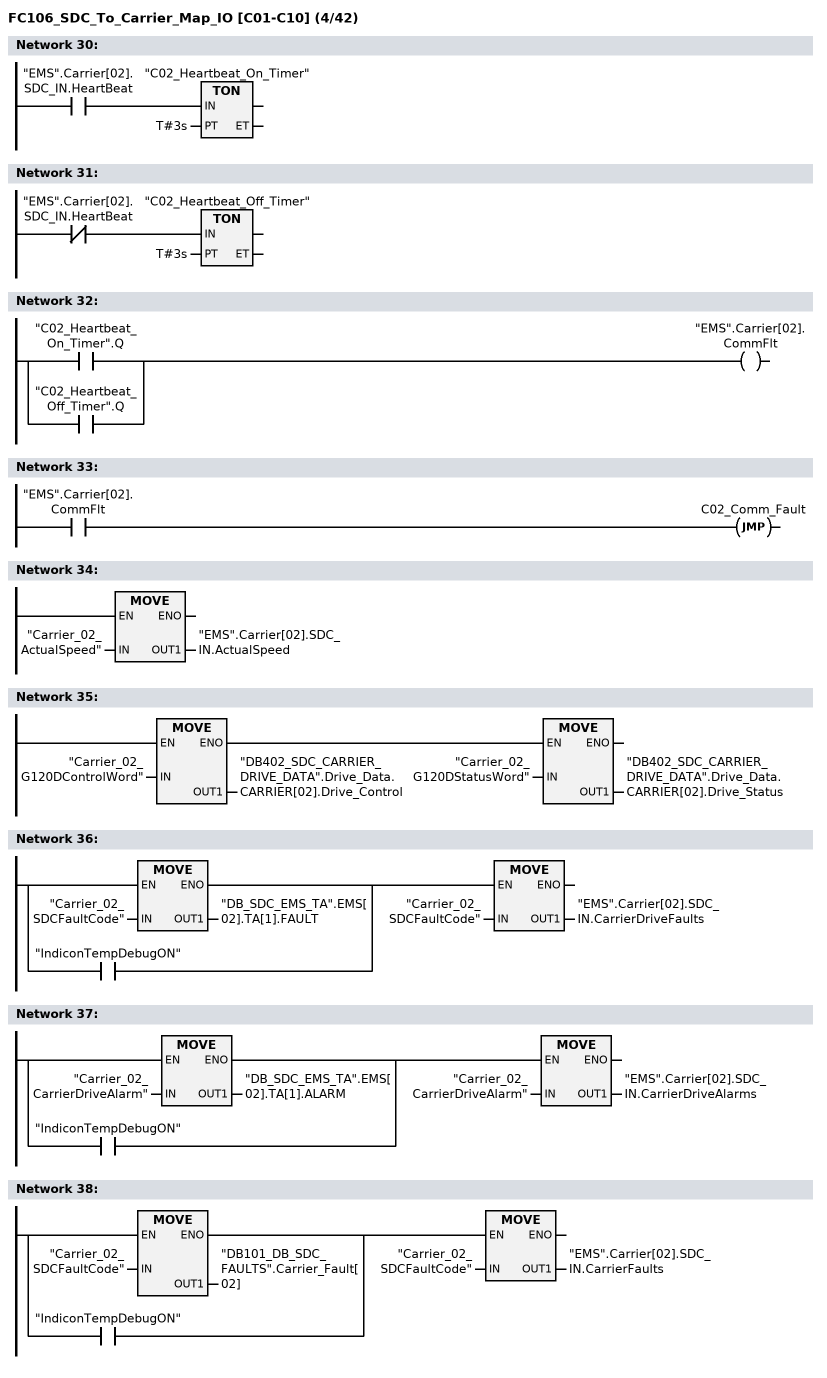
   "C02_Heartbeat_On_Timer".TON(IN := "EMS".Carrier[02].SDC_IN.HeartBeat, PT := T#3s);
END_REGION

REGION Network 31
   "C02_Heartbeat_Off_Timer".TON(IN := NOT "EMS".Carrier[02].SDC_IN.HeartBeat, PT := T#3s);
END_REGION

REGION Network 32
   RUNG wire#powerrail
      Contact( "C02_Heartbeat_On_Timer".Q )
      wire#w1
      Coil( "EMS".Carrier[02].CommFlt )
   END_RUNG
   RUNG wire#powerrail
      Contact( "C02_Heartbeat_Off_Timer".Q )
   END_RUNG wire#w1
   // the same network as SCL:
   "EMS".Carrier[02].CommFlt := "C02_Heartbeat_On_Timer".Q OR "C02_Heartbeat_Off_Timer".Q;
END_REGION

REGION Network 33
   RUNG wire#powerrail
      Contact( "EMS".Carrier[02].CommFlt )
      JumpCoil( C02_Comm_Fault )
   END_RUNG
   // the same network as SCL:
   IF "EMS".Carrier[02].CommFlt THEN GOTO C02_Comm_Fault; END_IF;
END_REGION

REGION Network 34
   RUNG wire#powerrail
      Move(in := "Carrier_02_ActualSpeed", out1 => "EMS".Carrier[02].SDC_IN.ActualSpeed)
   END_RUNG
   // the same network as SCL:
   "EMS".Carrier[02].SDC_IN.ActualSpeed := "Carrier_02_ActualSpeed";
END_REGION

REGION Network 35
   RUNG wire#powerrail
      Move(in := "Carrier_02_G120DControlWord", out1 => "DB402_SDC_CARRIER_DRIVE_DATA".Drive_Data.CARRIER[02].Drive_Control)
      Move(in := "Carrier_02_G120DStatusWord", out1 => "DB402_SDC_CARRIER_DRIVE_DATA".Drive_Data.CARRIER[02].Drive_Status)
   END_RUNG
   // the same network as SCL:
   "DB402_SDC_CARRIER_DRIVE_DATA".Drive_Data.CARRIER[02].Drive_Control := "Carrier_02_G120DControlWord";
   "DB402_SDC_CARRIER_DRIVE_DATA".Drive_Data.CARRIER[02].Drive_Status := "Carrier_02_G120DStatusWord";
END_REGION

REGION Network 36
   RUNG wire#powerrail
      Move(in := "Carrier_02_SDCFaultCode", out1 => "DB_SDC_EMS_TA".EMS[02].TA[1].FAULT)
      wire#w1
      Move(in := "Carrier_02_SDCFaultCode", out1 => "EMS".Carrier[02].SDC_IN.CarrierDriveFaults)
   END_RUNG
   RUNG wire#powerrail
      Contact( "IndiconTempDebugON" )
   END_RUNG wire#w1
   // the same network as SCL:
   "DB_SDC_EMS_TA".EMS[02].TA[1].FAULT := "Carrier_02_SDCFaultCode";
   IF TRUE OR "IndiconTempDebugON" THEN
       "EMS".Carrier[02].SDC_IN.CarrierDriveFaults := "Carrier_02_SDCFaultCode";
   END_IF;
END_REGION

REGION Network 37
   RUNG wire#powerrail
      Move(in := "Carrier_02_CarrierDriveAlarm", out1 => "DB_SDC_EMS_TA".EMS[02].TA[1].ALARM)
      wire#w1
      Move(in := "Carrier_02_CarrierDriveAlarm", out1 => "EMS".Carrier[02].SDC_IN.CarrierDriveAlarms)
   END_RUNG
   RUNG wire#powerrail
      Contact( "IndiconTempDebugON" )
   END_RUNG wire#w1
   // the same network as SCL:
   "DB_SDC_EMS_TA".EMS[02].TA[1].ALARM := "Carrier_02_CarrierDriveAlarm";
   IF TRUE OR "IndiconTempDebugON" THEN
       "EMS".Carrier[02].SDC_IN.CarrierDriveAlarms := "Carrier_02_CarrierDriveAlarm";
   END_IF;
END_REGION

REGION Network 38
   RUNG wire#powerrail
      Move(in := "Carrier_02_SDCFaultCode", out1 => "DB101_DB_SDC_FAULTS".Carrier_Fault[02])
      wire#w1
      Move(in := "Carrier_02_SDCFaultCode", out1 => "EMS".Carrier[02].SDC_IN.CarrierFaults)
   END_RUNG
   RUNG wire#powerrail
      Contact( "IndiconTempDebugON" )
   END_RUNG wire#w1
   // the same network as SCL:
   "DB101_DB_SDC_FAULTS".Carrier_Fault[02] := "Carrier_02_SDCFaultCode";
   IF TRUE OR "IndiconTempDebugON" THEN
       "EMS".Carrier[02].SDC_IN.CarrierFaults := "Carrier_02_SDCFaultCode";
   END_IF;
END_REGION

REGION Network 39
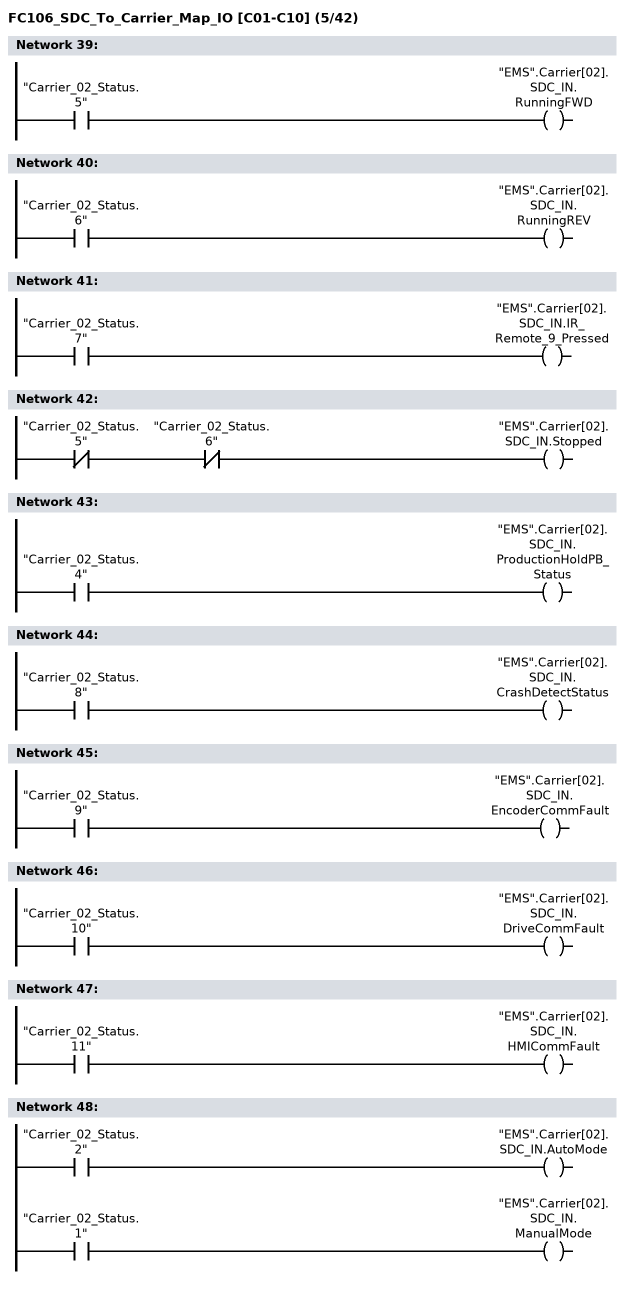
   RUNG wire#powerrail
      Contact( "Carrier_02_Status.5" )
      Coil( "EMS".Carrier[02].SDC_IN.RunningFWD )
   END_RUNG
   // the same network as SCL:
   "EMS".Carrier[02].SDC_IN.RunningFWD := "Carrier_02_Status.5";
END_REGION

REGION Network 40
   RUNG wire#powerrail
      Contact( "Carrier_02_Status.6" )
      Coil( "EMS".Carrier[02].SDC_IN.RunningREV )
   END_RUNG
   // the same network as SCL:
   "EMS".Carrier[02].SDC_IN.RunningREV := "Carrier_02_Status.6";
END_REGION

REGION Network 41
   RUNG wire#powerrail
      Contact( "Carrier_02_Status.7" )
      Coil( "EMS".Carrier[02].SDC_IN.IR_Remote_9_Pressed )
   END_RUNG
   // the same network as SCL:
   "EMS".Carrier[02].SDC_IN.IR_Remote_9_Pressed := "Carrier_02_Status.7";
END_REGION

REGION Network 42
   RUNG wire#powerrail
      I_Contact( "Carrier_02_Status.5" )
      I_Contact( "Carrier_02_Status.6" )
      Coil( "EMS".Carrier[02].SDC_IN.Stopped )
   END_RUNG
   // the same network as SCL:
   "EMS".Carrier[02].SDC_IN.Stopped := NOT "Carrier_02_Status.5" AND NOT "Carrier_02_Status.6";
END_REGION

REGION Network 43
   RUNG wire#powerrail
      Contact( "Carrier_02_Status.4" )
      Coil( "EMS".Carrier[02].SDC_IN.ProductionHoldPB_Status )
   END_RUNG
   // the same network as SCL:
   "EMS".Carrier[02].SDC_IN.ProductionHoldPB_Status := "Carrier_02_Status.4";
END_REGION

REGION Network 44
   RUNG wire#powerrail
      Contact( "Carrier_02_Status.8" )
      Coil( "EMS".Carrier[02].SDC_IN.CrashDetectStatus )
   END_RUNG
   // the same network as SCL:
   "EMS".Carrier[02].SDC_IN.CrashDetectStatus := "Carrier_02_Status.8";
END_REGION

REGION Network 45
   RUNG wire#powerrail
      Contact( "Carrier_02_Status.9" )
      Coil( "EMS".Carrier[02].SDC_IN.EncoderCommFault )
   END_RUNG
   // the same network as SCL:
   "EMS".Carrier[02].SDC_IN.EncoderCommFault := "Carrier_02_Status.9";
END_REGION

REGION Network 46
   RUNG wire#powerrail
      Contact( "Carrier_02_Status.10" )
      Coil( "EMS".Carrier[02].SDC_IN.DriveCommFault )
   END_RUNG
   // the same network as SCL:
   "EMS".Carrier[02].SDC_IN.DriveCommFault := "Carrier_02_Status.10";
END_REGION

REGION Network 47
   RUNG wire#powerrail
      Contact( "Carrier_02_Status.11" )
      Coil( "EMS".Carrier[02].SDC_IN.HMICommFault )
   END_RUNG
   // the same network as SCL:
   "EMS".Carrier[02].SDC_IN.HMICommFault := "Carrier_02_Status.11";
END_REGION

REGION Network 48
   RUNG wire#powerrail
      Contact( "Carrier_02_Status.2" )
      Coil( "EMS".Carrier[02].SDC_IN.AutoMode )
   END_RUNG
   RUNG wire#powerrail
      Contact( "Carrier_02_Status.1" )
      Coil( "EMS".Carrier[02].SDC_IN.ManualMode )
   END_RUNG
   // the same network as SCL:
   "EMS".Carrier[02].SDC_IN.AutoMode := "Carrier_02_Status.2";
   "EMS".Carrier[02].SDC_IN.ManualMode := "Carrier_02_Status.1";
END_REGION

REGION Network 49
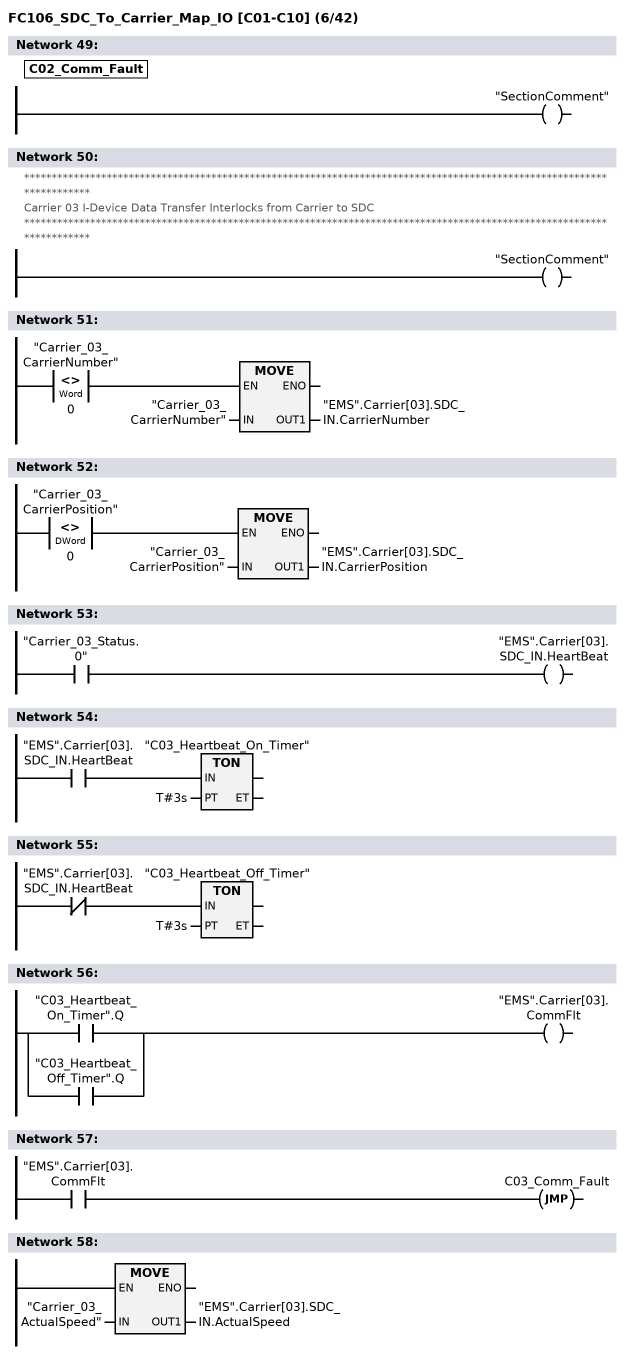
   Label( C02_Comm_Fault )
   RUNG wire#powerrail
      Coil( "SectionComment" )
   END_RUNG
   // the same network as SCL:
   C02_Comm_Fault:
   "SectionComment" := TRUE;
END_REGION

REGION Network 50
   // **********************************************************************************************************************
   // 
   // Carrier 03 I-Device Data Transfer Interlocks from Carrier to SDC
   // 
   // **********************************************************************************************************************
   RUNG wire#powerrail
      Coil( "SectionComment" )
   END_RUNG
   // the same network as SCL:
   "SectionComment" := TRUE;
END_REGION

REGION Network 51
   RUNG wire#powerrail
      { S7_Templates := "SrcType := Word" } NE_Contact(in1 := "Carrier_03_CarrierNumber", in2 := 0)
      Move(in := "Carrier_03_CarrierNumber", out1 => "EMS".Carrier[03].SDC_IN.CarrierNumber)
   END_RUNG
   // the same network as SCL:
   IF "Carrier_03_CarrierNumber" <> 0 THEN
       "EMS".Carrier[03].SDC_IN.CarrierNumber := "Carrier_03_CarrierNumber";
   END_IF;
END_REGION

REGION Network 52
   RUNG wire#powerrail
      { S7_Templates := "SrcType := DWord" } NE_Contact(in1 := "Carrier_03_CarrierPosition", in2 := 0)
      Move(in := "Carrier_03_CarrierPosition", out1 => "EMS".Carrier[03].SDC_IN.CarrierPosition)
   END_RUNG
   // the same network as SCL:
   IF "Carrier_03_CarrierPosition" <> 0 THEN
       "EMS".Carrier[03].SDC_IN.CarrierPosition := "Carrier_03_CarrierPosition";
   END_IF;
END_REGION

REGION Network 53
   RUNG wire#powerrail
      Contact( "Carrier_03_Status.0" )
      Coil( "EMS".Carrier[03].SDC_IN.HeartBeat )
   END_RUNG
   // the same network as SCL:
   "EMS".Carrier[03].SDC_IN.HeartBeat := "Carrier_03_Status.0";
END_REGION

REGION Network 54
   "C03_Heartbeat_On_Timer".TON(IN := "EMS".Carrier[03].SDC_IN.HeartBeat, PT := T#3s);
END_REGION

REGION Network 55
   "C03_Heartbeat_Off_Timer".TON(IN := NOT "EMS".Carrier[03].SDC_IN.HeartBeat, PT := T#3s);
END_REGION

REGION Network 56
   RUNG wire#powerrail
      Contact( "C03_Heartbeat_On_Timer".Q )
      wire#w1
      Coil( "EMS".Carrier[03].CommFlt )
   END_RUNG
   RUNG wire#powerrail
      Contact( "C03_Heartbeat_Off_Timer".Q )
   END_RUNG wire#w1
   // the same network as SCL:
   "EMS".Carrier[03].CommFlt := "C03_Heartbeat_On_Timer".Q OR "C03_Heartbeat_Off_Timer".Q;
END_REGION

REGION Network 57
   RUNG wire#powerrail
      Contact( "EMS".Carrier[03].CommFlt )
      JumpCoil( C03_Comm_Fault )
   END_RUNG
   // the same network as SCL:
   IF "EMS".Carrier[03].CommFlt THEN GOTO C03_Comm_Fault; END_IF;
END_REGION

REGION Network 58
   RUNG wire#powerrail
      Move(in := "Carrier_03_ActualSpeed", out1 => "EMS".Carrier[03].SDC_IN.ActualSpeed)
   END_RUNG
   // the same network as SCL:
   "EMS".Carrier[03].SDC_IN.ActualSpeed := "Carrier_03_ActualSpeed";
END_REGION

REGION Network 59
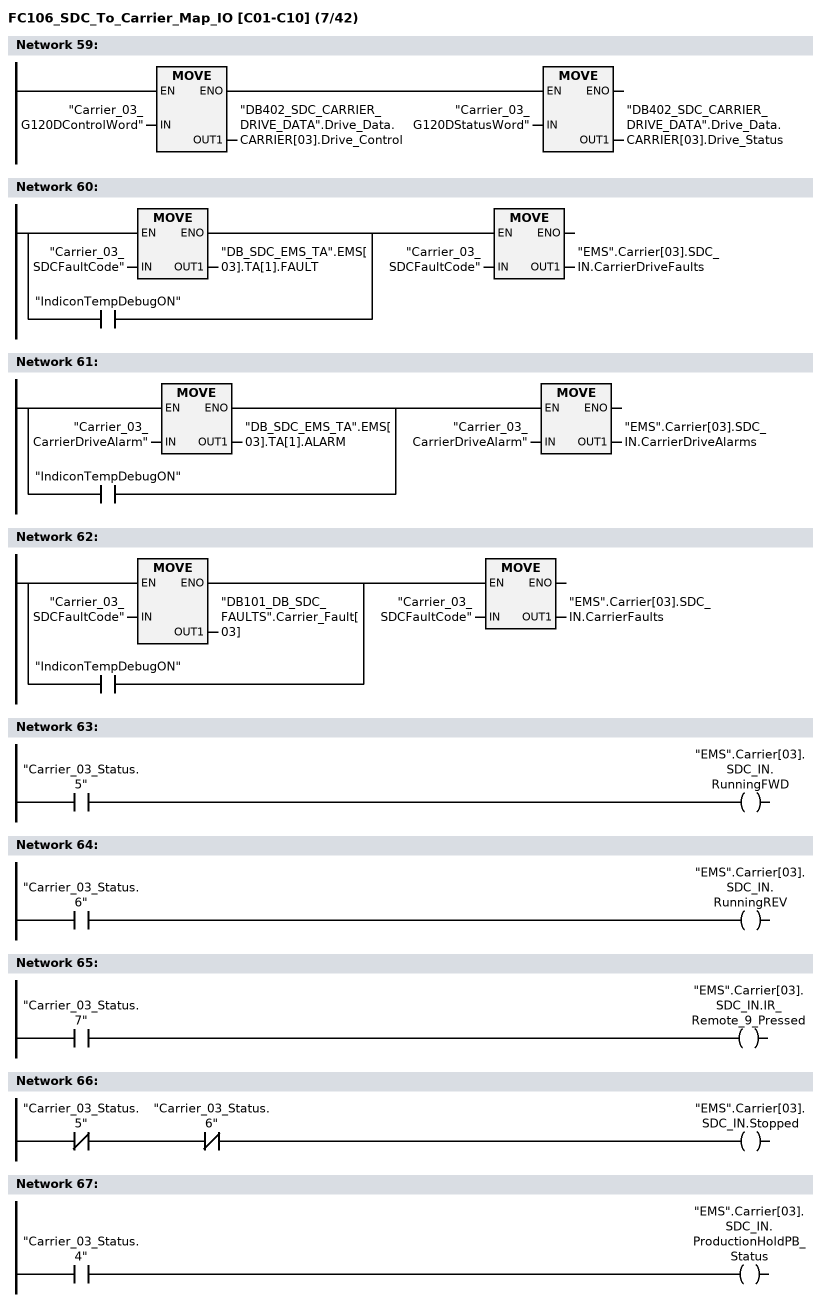
   RUNG wire#powerrail
      Move(in := "Carrier_03_G120DControlWord", out1 => "DB402_SDC_CARRIER_DRIVE_DATA".Drive_Data.CARRIER[03].Drive_Control)
      Move(in := "Carrier_03_G120DStatusWord", out1 => "DB402_SDC_CARRIER_DRIVE_DATA".Drive_Data.CARRIER[03].Drive_Status)
   END_RUNG
   // the same network as SCL:
   "DB402_SDC_CARRIER_DRIVE_DATA".Drive_Data.CARRIER[03].Drive_Control := "Carrier_03_G120DControlWord";
   "DB402_SDC_CARRIER_DRIVE_DATA".Drive_Data.CARRIER[03].Drive_Status := "Carrier_03_G120DStatusWord";
END_REGION

REGION Network 60
   RUNG wire#powerrail
      Move(in := "Carrier_03_SDCFaultCode", out1 => "DB_SDC_EMS_TA".EMS[03].TA[1].FAULT)
      wire#w1
      Move(in := "Carrier_03_SDCFaultCode", out1 => "EMS".Carrier[03].SDC_IN.CarrierDriveFaults)
   END_RUNG
   RUNG wire#powerrail
      Contact( "IndiconTempDebugON" )
   END_RUNG wire#w1
   // the same network as SCL:
   "DB_SDC_EMS_TA".EMS[03].TA[1].FAULT := "Carrier_03_SDCFaultCode";
   IF TRUE OR "IndiconTempDebugON" THEN
       "EMS".Carrier[03].SDC_IN.CarrierDriveFaults := "Carrier_03_SDCFaultCode";
   END_IF;
END_REGION

REGION Network 61
   RUNG wire#powerrail
      Move(in := "Carrier_03_CarrierDriveAlarm", out1 => "DB_SDC_EMS_TA".EMS[03].TA[1].ALARM)
      wire#w1
      Move(in := "Carrier_03_CarrierDriveAlarm", out1 => "EMS".Carrier[03].SDC_IN.CarrierDriveAlarms)
   END_RUNG
   RUNG wire#powerrail
      Contact( "IndiconTempDebugON" )
   END_RUNG wire#w1
   // the same network as SCL:
   "DB_SDC_EMS_TA".EMS[03].TA[1].ALARM := "Carrier_03_CarrierDriveAlarm";
   IF TRUE OR "IndiconTempDebugON" THEN
       "EMS".Carrier[03].SDC_IN.CarrierDriveAlarms := "Carrier_03_CarrierDriveAlarm";
   END_IF;
END_REGION

REGION Network 62
   RUNG wire#powerrail
      Move(in := "Carrier_03_SDCFaultCode", out1 => "DB101_DB_SDC_FAULTS".Carrier_Fault[03])
      wire#w1
      Move(in := "Carrier_03_SDCFaultCode", out1 => "EMS".Carrier[03].SDC_IN.CarrierFaults)
   END_RUNG
   RUNG wire#powerrail
      Contact( "IndiconTempDebugON" )
   END_RUNG wire#w1
   // the same network as SCL:
   "DB101_DB_SDC_FAULTS".Carrier_Fault[03] := "Carrier_03_SDCFaultCode";
   IF TRUE OR "IndiconTempDebugON" THEN
       "EMS".Carrier[03].SDC_IN.CarrierFaults := "Carrier_03_SDCFaultCode";
   END_IF;
END_REGION

REGION Network 63
   RUNG wire#powerrail
      Contact( "Carrier_03_Status.5" )
      Coil( "EMS".Carrier[03].SDC_IN.RunningFWD )
   END_RUNG
   // the same network as SCL:
   "EMS".Carrier[03].SDC_IN.RunningFWD := "Carrier_03_Status.5";
END_REGION

REGION Network 64
   RUNG wire#powerrail
      Contact( "Carrier_03_Status.6" )
      Coil( "EMS".Carrier[03].SDC_IN.RunningREV )
   END_RUNG
   // the same network as SCL:
   "EMS".Carrier[03].SDC_IN.RunningREV := "Carrier_03_Status.6";
END_REGION

REGION Network 65
   RUNG wire#powerrail
      Contact( "Carrier_03_Status.7" )
      Coil( "EMS".Carrier[03].SDC_IN.IR_Remote_9_Pressed )
   END_RUNG
   // the same network as SCL:
   "EMS".Carrier[03].SDC_IN.IR_Remote_9_Pressed := "Carrier_03_Status.7";
END_REGION

REGION Network 66
   RUNG wire#powerrail
      I_Contact( "Carrier_03_Status.5" )
      I_Contact( "Carrier_03_Status.6" )
      Coil( "EMS".Carrier[03].SDC_IN.Stopped )
   END_RUNG
   // the same network as SCL:
   "EMS".Carrier[03].SDC_IN.Stopped := NOT "Carrier_03_Status.5" AND NOT "Carrier_03_Status.6";
END_REGION

REGION Network 67
   RUNG wire#powerrail
      Contact( "Carrier_03_Status.4" )
      Coil( "EMS".Carrier[03].SDC_IN.ProductionHoldPB_Status )
   END_RUNG
   // the same network as SCL:
   "EMS".Carrier[03].SDC_IN.ProductionHoldPB_Status := "Carrier_03_Status.4";
END_REGION

REGION Network 68
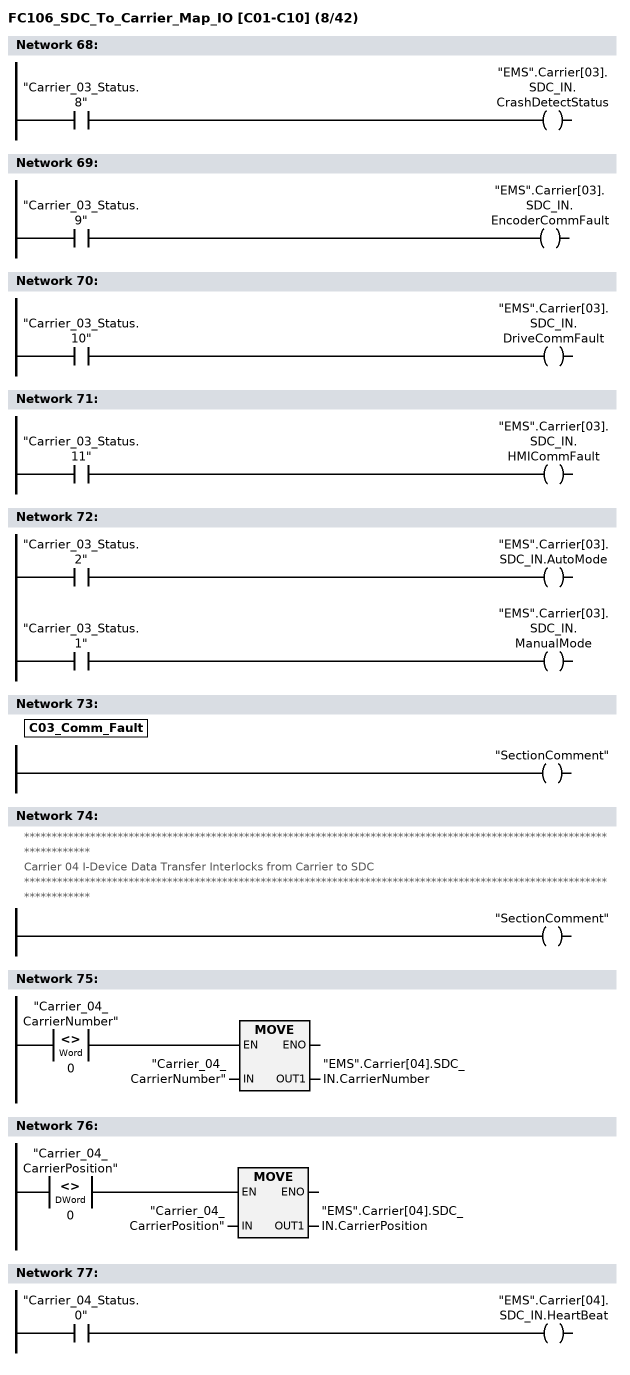
   RUNG wire#powerrail
      Contact( "Carrier_03_Status.8" )
      Coil( "EMS".Carrier[03].SDC_IN.CrashDetectStatus )
   END_RUNG
   // the same network as SCL:
   "EMS".Carrier[03].SDC_IN.CrashDetectStatus := "Carrier_03_Status.8";
END_REGION

REGION Network 69
   RUNG wire#powerrail
      Contact( "Carrier_03_Status.9" )
      Coil( "EMS".Carrier[03].SDC_IN.EncoderCommFault )
   END_RUNG
   // the same network as SCL:
   "EMS".Carrier[03].SDC_IN.EncoderCommFault := "Carrier_03_Status.9";
END_REGION

REGION Network 70
   RUNG wire#powerrail
      Contact( "Carrier_03_Status.10" )
      Coil( "EMS".Carrier[03].SDC_IN.DriveCommFault )
   END_RUNG
   // the same network as SCL:
   "EMS".Carrier[03].SDC_IN.DriveCommFault := "Carrier_03_Status.10";
END_REGION

REGION Network 71
   RUNG wire#powerrail
      Contact( "Carrier_03_Status.11" )
      Coil( "EMS".Carrier[03].SDC_IN.HMICommFault )
   END_RUNG
   // the same network as SCL:
   "EMS".Carrier[03].SDC_IN.HMICommFault := "Carrier_03_Status.11";
END_REGION

REGION Network 72
   RUNG wire#powerrail
      Contact( "Carrier_03_Status.2" )
      Coil( "EMS".Carrier[03].SDC_IN.AutoMode )
   END_RUNG
   RUNG wire#powerrail
      Contact( "Carrier_03_Status.1" )
      Coil( "EMS".Carrier[03].SDC_IN.ManualMode )
   END_RUNG
   // the same network as SCL:
   "EMS".Carrier[03].SDC_IN.AutoMode := "Carrier_03_Status.2";
   "EMS".Carrier[03].SDC_IN.ManualMode := "Carrier_03_Status.1";
END_REGION

REGION Network 73
   Label( C03_Comm_Fault )
   RUNG wire#powerrail
      Coil( "SectionComment" )
   END_RUNG
   // the same network as SCL:
   C03_Comm_Fault:
   "SectionComment" := TRUE;
END_REGION

REGION Network 74
   // **********************************************************************************************************************
   // 
   // Carrier 04 I-Device Data Transfer Interlocks from Carrier to SDC
   // 
   // **********************************************************************************************************************
   RUNG wire#powerrail
      Coil( "SectionComment" )
   END_RUNG
   // the same network as SCL:
   "SectionComment" := TRUE;
END_REGION

REGION Network 75
   RUNG wire#powerrail
      { S7_Templates := "SrcType := Word" } NE_Contact(in1 := "Carrier_04_CarrierNumber", in2 := 0)
      Move(in := "Carrier_04_CarrierNumber", out1 => "EMS".Carrier[04].SDC_IN.CarrierNumber)
   END_RUNG
   // the same network as SCL:
   IF "Carrier_04_CarrierNumber" <> 0 THEN
       "EMS".Carrier[04].SDC_IN.CarrierNumber := "Carrier_04_CarrierNumber";
   END_IF;
END_REGION

REGION Network 76
   RUNG wire#powerrail
      { S7_Templates := "SrcType := DWord" } NE_Contact(in1 := "Carrier_04_CarrierPosition", in2 := 0)
      Move(in := "Carrier_04_CarrierPosition", out1 => "EMS".Carrier[04].SDC_IN.CarrierPosition)
   END_RUNG
   // the same network as SCL:
   IF "Carrier_04_CarrierPosition" <> 0 THEN
       "EMS".Carrier[04].SDC_IN.CarrierPosition := "Carrier_04_CarrierPosition";
   END_IF;
END_REGION

REGION Network 77
   RUNG wire#powerrail
      Contact( "Carrier_04_Status.0" )
      Coil( "EMS".Carrier[04].SDC_IN.HeartBeat )
   END_RUNG
   // the same network as SCL:
   "EMS".Carrier[04].SDC_IN.HeartBeat := "Carrier_04_Status.0";
END_REGION

REGION Network 78
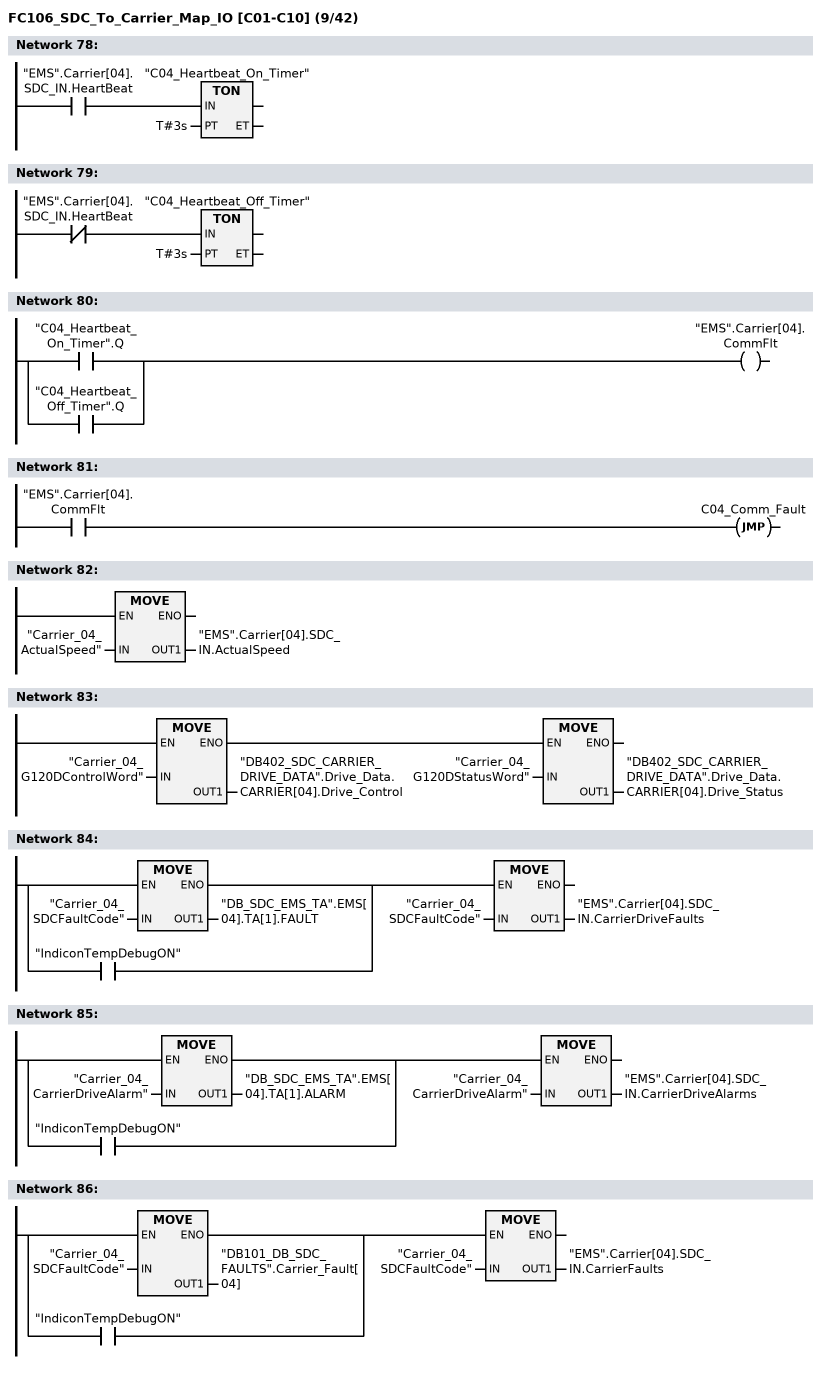
   "C04_Heartbeat_On_Timer".TON(IN := "EMS".Carrier[04].SDC_IN.HeartBeat, PT := T#3s);
END_REGION

REGION Network 79
   "C04_Heartbeat_Off_Timer".TON(IN := NOT "EMS".Carrier[04].SDC_IN.HeartBeat, PT := T#3s);
END_REGION

REGION Network 80
   RUNG wire#powerrail
      Contact( "C04_Heartbeat_On_Timer".Q )
      wire#w1
      Coil( "EMS".Carrier[04].CommFlt )
   END_RUNG
   RUNG wire#powerrail
      Contact( "C04_Heartbeat_Off_Timer".Q )
   END_RUNG wire#w1
   // the same network as SCL:
   "EMS".Carrier[04].CommFlt := "C04_Heartbeat_On_Timer".Q OR "C04_Heartbeat_Off_Timer".Q;
END_REGION

REGION Network 81
   RUNG wire#powerrail
      Contact( "EMS".Carrier[04].CommFlt )
      JumpCoil( C04_Comm_Fault )
   END_RUNG
   // the same network as SCL:
   IF "EMS".Carrier[04].CommFlt THEN GOTO C04_Comm_Fault; END_IF;
END_REGION

REGION Network 82
   RUNG wire#powerrail
      Move(in := "Carrier_04_ActualSpeed", out1 => "EMS".Carrier[04].SDC_IN.ActualSpeed)
   END_RUNG
   // the same network as SCL:
   "EMS".Carrier[04].SDC_IN.ActualSpeed := "Carrier_04_ActualSpeed";
END_REGION

REGION Network 83
   RUNG wire#powerrail
      Move(in := "Carrier_04_G120DControlWord", out1 => "DB402_SDC_CARRIER_DRIVE_DATA".Drive_Data.CARRIER[04].Drive_Control)
      Move(in := "Carrier_04_G120DStatusWord", out1 => "DB402_SDC_CARRIER_DRIVE_DATA".Drive_Data.CARRIER[04].Drive_Status)
   END_RUNG
   // the same network as SCL:
   "DB402_SDC_CARRIER_DRIVE_DATA".Drive_Data.CARRIER[04].Drive_Control := "Carrier_04_G120DControlWord";
   "DB402_SDC_CARRIER_DRIVE_DATA".Drive_Data.CARRIER[04].Drive_Status := "Carrier_04_G120DStatusWord";
END_REGION

REGION Network 84
   RUNG wire#powerrail
      Move(in := "Carrier_04_SDCFaultCode", out1 => "DB_SDC_EMS_TA".EMS[04].TA[1].FAULT)
      wire#w1
      Move(in := "Carrier_04_SDCFaultCode", out1 => "EMS".Carrier[04].SDC_IN.CarrierDriveFaults)
   END_RUNG
   RUNG wire#powerrail
      Contact( "IndiconTempDebugON" )
   END_RUNG wire#w1
   // the same network as SCL:
   "DB_SDC_EMS_TA".EMS[04].TA[1].FAULT := "Carrier_04_SDCFaultCode";
   IF TRUE OR "IndiconTempDebugON" THEN
       "EMS".Carrier[04].SDC_IN.CarrierDriveFaults := "Carrier_04_SDCFaultCode";
   END_IF;
END_REGION

REGION Network 85
   RUNG wire#powerrail
      Move(in := "Carrier_04_CarrierDriveAlarm", out1 => "DB_SDC_EMS_TA".EMS[04].TA[1].ALARM)
      wire#w1
      Move(in := "Carrier_04_CarrierDriveAlarm", out1 => "EMS".Carrier[04].SDC_IN.CarrierDriveAlarms)
   END_RUNG
   RUNG wire#powerrail
      Contact( "IndiconTempDebugON" )
   END_RUNG wire#w1
   // the same network as SCL:
   "DB_SDC_EMS_TA".EMS[04].TA[1].ALARM := "Carrier_04_CarrierDriveAlarm";
   IF TRUE OR "IndiconTempDebugON" THEN
       "EMS".Carrier[04].SDC_IN.CarrierDriveAlarms := "Carrier_04_CarrierDriveAlarm";
   END_IF;
END_REGION

REGION Network 86
   RUNG wire#powerrail
      Move(in := "Carrier_04_SDCFaultCode", out1 => "DB101_DB_SDC_FAULTS".Carrier_Fault[04])
      wire#w1
      Move(in := "Carrier_04_SDCFaultCode", out1 => "EMS".Carrier[04].SDC_IN.CarrierFaults)
   END_RUNG
   RUNG wire#powerrail
      Contact( "IndiconTempDebugON" )
   END_RUNG wire#w1
   // the same network as SCL:
   "DB101_DB_SDC_FAULTS".Carrier_Fault[04] := "Carrier_04_SDCFaultCode";
   IF TRUE OR "IndiconTempDebugON" THEN
       "EMS".Carrier[04].SDC_IN.CarrierFaults := "Carrier_04_SDCFaultCode";
   END_IF;
END_REGION

REGION Network 87
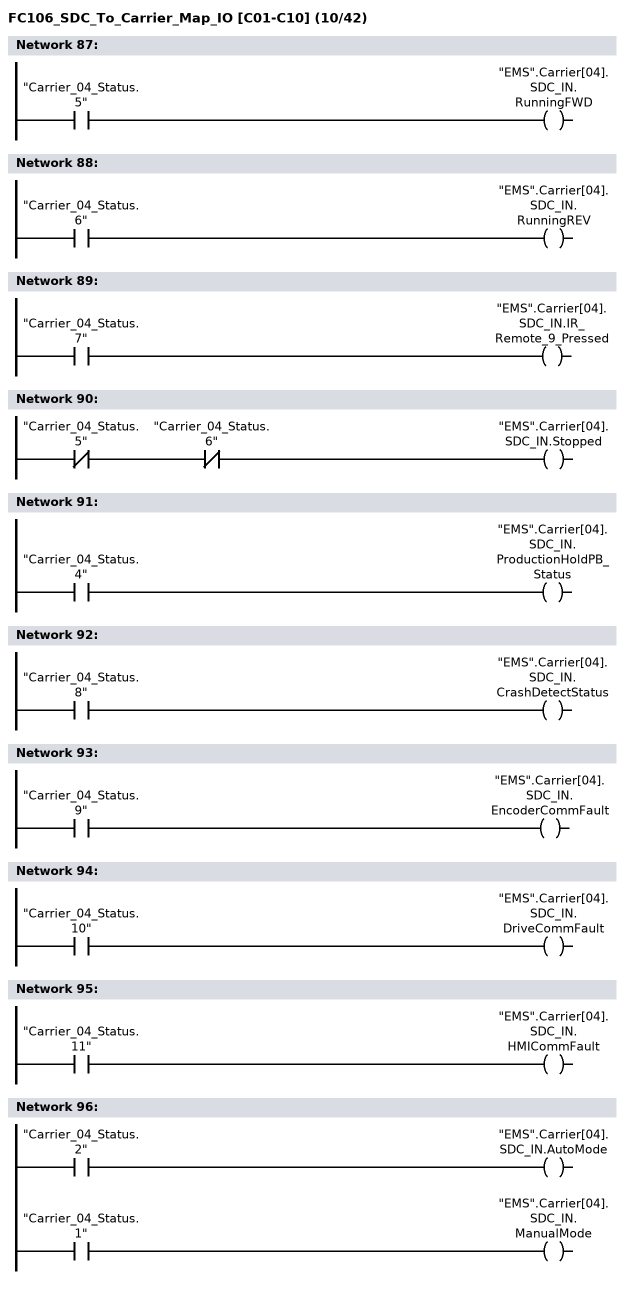
   RUNG wire#powerrail
      Contact( "Carrier_04_Status.5" )
      Coil( "EMS".Carrier[04].SDC_IN.RunningFWD )
   END_RUNG
   // the same network as SCL:
   "EMS".Carrier[04].SDC_IN.RunningFWD := "Carrier_04_Status.5";
END_REGION

REGION Network 88
   RUNG wire#powerrail
      Contact( "Carrier_04_Status.6" )
      Coil( "EMS".Carrier[04].SDC_IN.RunningREV )
   END_RUNG
   // the same network as SCL:
   "EMS".Carrier[04].SDC_IN.RunningREV := "Carrier_04_Status.6";
END_REGION

REGION Network 89
   RUNG wire#powerrail
      Contact( "Carrier_04_Status.7" )
      Coil( "EMS".Carrier[04].SDC_IN.IR_Remote_9_Pressed )
   END_RUNG
   // the same network as SCL:
   "EMS".Carrier[04].SDC_IN.IR_Remote_9_Pressed := "Carrier_04_Status.7";
END_REGION

REGION Network 90
   RUNG wire#powerrail
      I_Contact( "Carrier_04_Status.5" )
      I_Contact( "Carrier_04_Status.6" )
      Coil( "EMS".Carrier[04].SDC_IN.Stopped )
   END_RUNG
   // the same network as SCL:
   "EMS".Carrier[04].SDC_IN.Stopped := NOT "Carrier_04_Status.5" AND NOT "Carrier_04_Status.6";
END_REGION

REGION Network 91
   RUNG wire#powerrail
      Contact( "Carrier_04_Status.4" )
      Coil( "EMS".Carrier[04].SDC_IN.ProductionHoldPB_Status )
   END_RUNG
   // the same network as SCL:
   "EMS".Carrier[04].SDC_IN.ProductionHoldPB_Status := "Carrier_04_Status.4";
END_REGION

REGION Network 92
   RUNG wire#powerrail
      Contact( "Carrier_04_Status.8" )
      Coil( "EMS".Carrier[04].SDC_IN.CrashDetectStatus )
   END_RUNG
   // the same network as SCL:
   "EMS".Carrier[04].SDC_IN.CrashDetectStatus := "Carrier_04_Status.8";
END_REGION

REGION Network 93
   RUNG wire#powerrail
      Contact( "Carrier_04_Status.9" )
      Coil( "EMS".Carrier[04].SDC_IN.EncoderCommFault )
   END_RUNG
   // the same network as SCL:
   "EMS".Carrier[04].SDC_IN.EncoderCommFault := "Carrier_04_Status.9";
END_REGION

REGION Network 94
   RUNG wire#powerrail
      Contact( "Carrier_04_Status.10" )
      Coil( "EMS".Carrier[04].SDC_IN.DriveCommFault )
   END_RUNG
   // the same network as SCL:
   "EMS".Carrier[04].SDC_IN.DriveCommFault := "Carrier_04_Status.10";
END_REGION

REGION Network 95
   RUNG wire#powerrail
      Contact( "Carrier_04_Status.11" )
      Coil( "EMS".Carrier[04].SDC_IN.HMICommFault )
   END_RUNG
   // the same network as SCL:
   "EMS".Carrier[04].SDC_IN.HMICommFault := "Carrier_04_Status.11";
END_REGION

REGION Network 96
   RUNG wire#powerrail
      Contact( "Carrier_04_Status.2" )
      Coil( "EMS".Carrier[04].SDC_IN.AutoMode )
   END_RUNG
   RUNG wire#powerrail
      Contact( "Carrier_04_Status.1" )
      Coil( "EMS".Carrier[04].SDC_IN.ManualMode )
   END_RUNG
   // the same network as SCL:
   "EMS".Carrier[04].SDC_IN.AutoMode := "Carrier_04_Status.2";
   "EMS".Carrier[04].SDC_IN.ManualMode := "Carrier_04_Status.1";
END_REGION

REGION Network 97
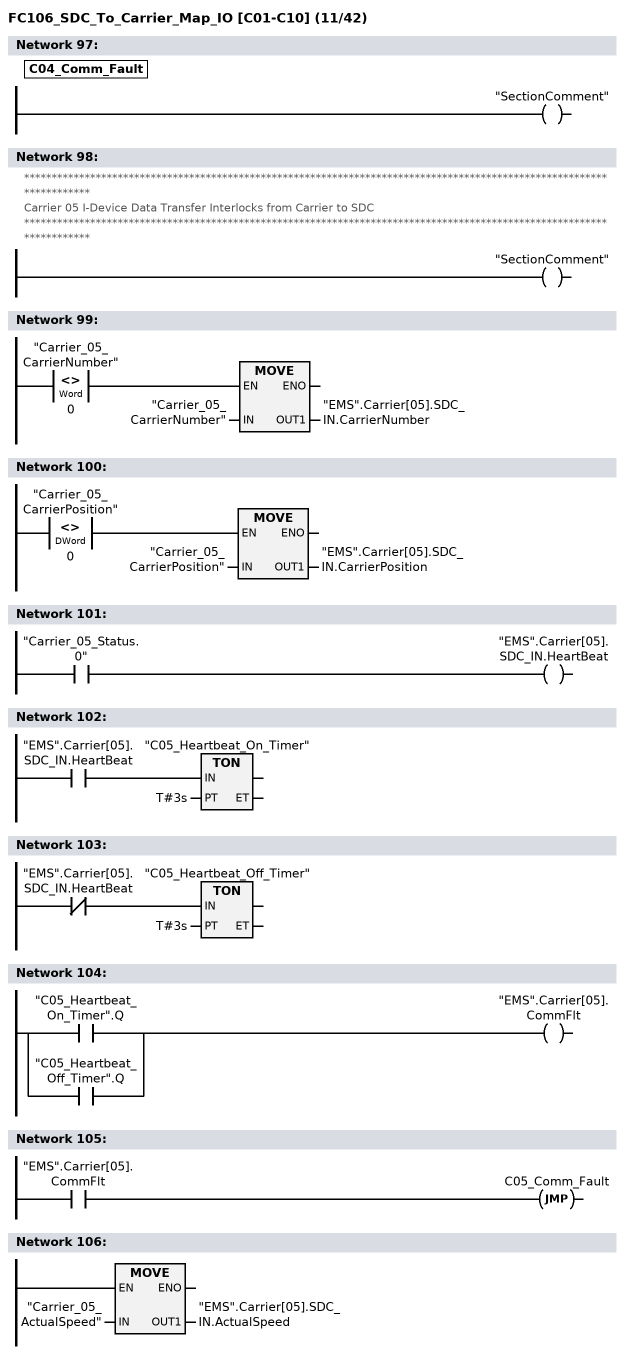
   Label( C04_Comm_Fault )
   RUNG wire#powerrail
      Coil( "SectionComment" )
   END_RUNG
   // the same network as SCL:
   C04_Comm_Fault:
   "SectionComment" := TRUE;
END_REGION

REGION Network 98
   // **********************************************************************************************************************
   // 
   // Carrier 05 I-Device Data Transfer Interlocks from Carrier to SDC
   // 
   // **********************************************************************************************************************
   RUNG wire#powerrail
      Coil( "SectionComment" )
   END_RUNG
   // the same network as SCL:
   "SectionComment" := TRUE;
END_REGION

REGION Network 99
   RUNG wire#powerrail
      { S7_Templates := "SrcType := Word" } NE_Contact(in1 := "Carrier_05_CarrierNumber", in2 := 0)
      Move(in := "Carrier_05_CarrierNumber", out1 => "EMS".Carrier[05].SDC_IN.CarrierNumber)
   END_RUNG
   // the same network as SCL:
   IF "Carrier_05_CarrierNumber" <> 0 THEN
       "EMS".Carrier[05].SDC_IN.CarrierNumber := "Carrier_05_CarrierNumber";
   END_IF;
END_REGION

REGION Network 100
   RUNG wire#powerrail
      { S7_Templates := "SrcType := DWord" } NE_Contact(in1 := "Carrier_05_CarrierPosition", in2 := 0)
      Move(in := "Carrier_05_CarrierPosition", out1 => "EMS".Carrier[05].SDC_IN.CarrierPosition)
   END_RUNG
   // the same network as SCL:
   IF "Carrier_05_CarrierPosition" <> 0 THEN
       "EMS".Carrier[05].SDC_IN.CarrierPosition := "Carrier_05_CarrierPosition";
   END_IF;
END_REGION

REGION Network 101
   RUNG wire#powerrail
      Contact( "Carrier_05_Status.0" )
      Coil( "EMS".Carrier[05].SDC_IN.HeartBeat )
   END_RUNG
   // the same network as SCL:
   "EMS".Carrier[05].SDC_IN.HeartBeat := "Carrier_05_Status.0";
END_REGION

REGION Network 102
   "C05_Heartbeat_On_Timer".TON(IN := "EMS".Carrier[05].SDC_IN.HeartBeat, PT := T#3s);
END_REGION

REGION Network 103
   "C05_Heartbeat_Off_Timer".TON(IN := NOT "EMS".Carrier[05].SDC_IN.HeartBeat, PT := T#3s);
END_REGION

REGION Network 104
   RUNG wire#powerrail
      Contact( "C05_Heartbeat_On_Timer".Q )
      wire#w1
      Coil( "EMS".Carrier[05].CommFlt )
   END_RUNG
   RUNG wire#powerrail
      Contact( "C05_Heartbeat_Off_Timer".Q )
   END_RUNG wire#w1
   // the same network as SCL:
   "EMS".Carrier[05].CommFlt := "C05_Heartbeat_On_Timer".Q OR "C05_Heartbeat_Off_Timer".Q;
END_REGION

REGION Network 105
   RUNG wire#powerrail
      Contact( "EMS".Carrier[05].CommFlt )
      JumpCoil( C05_Comm_Fault )
   END_RUNG
   // the same network as SCL:
   IF "EMS".Carrier[05].CommFlt THEN GOTO C05_Comm_Fault; END_IF;
END_REGION

REGION Network 106
   RUNG wire#powerrail
      Move(in := "Carrier_05_ActualSpeed", out1 => "EMS".Carrier[05].SDC_IN.ActualSpeed)
   END_RUNG
   // the same network as SCL:
   "EMS".Carrier[05].SDC_IN.ActualSpeed := "Carrier_05_ActualSpeed";
END_REGION

REGION Network 107
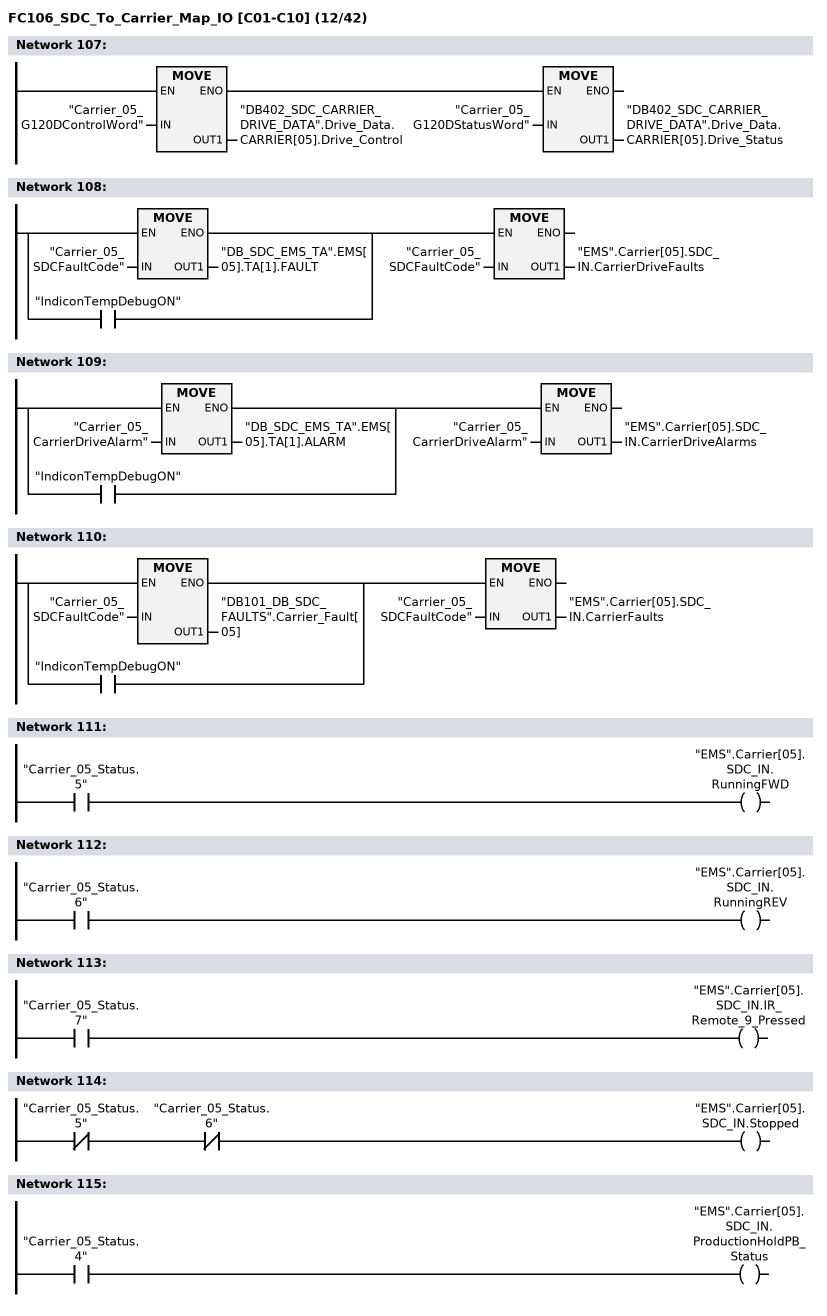
   RUNG wire#powerrail
      Move(in := "Carrier_05_G120DControlWord", out1 => "DB402_SDC_CARRIER_DRIVE_DATA".Drive_Data.CARRIER[05].Drive_Control)
      Move(in := "Carrier_05_G120DStatusWord", out1 => "DB402_SDC_CARRIER_DRIVE_DATA".Drive_Data.CARRIER[05].Drive_Status)
   END_RUNG
   // the same network as SCL:
   "DB402_SDC_CARRIER_DRIVE_DATA".Drive_Data.CARRIER[05].Drive_Control := "Carrier_05_G120DControlWord";
   "DB402_SDC_CARRIER_DRIVE_DATA".Drive_Data.CARRIER[05].Drive_Status := "Carrier_05_G120DStatusWord";
END_REGION
